TYPE "UDT_Actions"
VERSION : 0.1
   STRUCT
      MCMovement01WP : Bool;   // 1: Fapo in Vorpos AS
      MCMovement02WP : Bool;   // 2: Fapo in AS
      MCMovement03WP : Bool;   // 3: Fapu in Vorpos AS
      MCMovement04WP : Bool;   // 4: Fapu in AS
      MCMovement05WP : Bool;   // 5: Gestell in Vorpos AS
      MCMovement06WP : Bool;   // 6: Gestell in AS
      MCMovement07WP : Bool;   // 7: Parallelhub in Vorpos AS
      MCMovement08WP : Bool;   // 8: Parallelhub in AS
      MCMovement09WP : Bool;   // 9: Parallelhub unten (Fapu mit Fapo) verriegeln
      MCMovement10WP : Bool;   // 10: Sicherheitsriegel Parallelhub entriegeln
      MCMovement11WP : Bool;   // 11: Luftkissen aufblasen
      MCMovement12WP : Bool;   // 12: Form erkannt
      MCMovement13WP : Bool;   // 13: Sicherheitsriegel Fapo entriegeln
      MCMovement14WP : Bool;   // 14: Fapo referenzieren
      MCMovement15WP : Bool;   // 15: Fapu referenzieren
      MCMovement16WP : Bool;   // 16: Gestell referenzieren
      MCMovement17WP : Bool;   // 17: Rolltor zu
      MCMovement18WP : Bool;   // 18: Anschlag Fapo verriegeln
      MCMovement19WP : Bool;   // 19: Sicherheitsriegel Gestell entriegeln
      MCMovement20WP : Bool;   // 20:
      MCMovement21WP : Bool;   // 21:
      MCMovement22WP : Bool;   // 22:
      MCMovement23WP : Bool;   // 23:
      MCMovement24WP : Bool;   // 24:
      MCMovement25WP : Bool;   // 25: Werkzeugriegel Fapo verriegeln
      MCMovement26WP : Bool;   // 26: Werkzeugriegel Fapu verriegeln
      MCMovement27WP : Bool;   // 27: Hubleiste Fapu absenken
      MCMovement28WP : Bool;   // 28: Luftkissen aufblasen (kleiner Druck für Magnet)
      MCMovement29WP : Bool;   // 29: Magnetplatte Fapo einschalten
      MCMovement30WP : Bool;   // 30: Magnetplatte Fapu einschalten
      MCMovement31WP : Bool;   // 31: Fallsicherung Fapo verriegeln
      MCMovement32WP : Bool;   // 32: Fallsicherung Fapu verriegeln
      MCMovement01BP : Bool;   // 33: Fapo in Vorpos GS
      MCMovement02BP : Bool;   // 34: Fapo in GS
      MCMovement03BP : Bool;   // 35: Fapu in Vorpos GS
      MCMovement04BP : Bool;   // 36: Fapu in GS
      MCMovement05BP : Bool;   // 37: Gestell in Vorpos GS
      MCMovement06BP : Bool;   // 38: Gestell in GS
      MCMovement07BP : Bool;   // 39: Parallelhub in Vorpos GS
      MCMovement08BP : Bool;   // 40: Parallelhub in GS
      MCMovement09BP : Bool;   // 41: Parallelhub unten (Fapu mit Fapo) entriegeln
      MCMovement10BP : Bool;   // 42: Sicherheitsriegel Parallelhub verriegeln
      MCMovement11BP : Bool;   // 43: Luftkissen ablassen
      MCMovement12BP : Bool;   // 44:
      MCMovement13BP : Bool;   // 45: Sicherheitsriegel Fapo verriegeln
      MCMovement14BP : Bool;   // 46: Parallelhub in GS od. in Vorpos GS
      MCMovement15BP : Bool;   // 47:
      MCMovement16BP : Bool;   // 48: Parallelhub referenzieren
      MCMovement17BP : Bool;   // 49: Rolltor auf
      MCMovement18BP : Bool;   // 50: Anschlag Fapo entriegeln
      MCMovement19BP : Bool;   // 51: Sicherheitsriegel Gestell verriegeln
      MCMovement20BP : Bool;   // 52:
      MCMovement21BP : Bool;   // 53:
      MCMovement22BP : Bool;   // 54:
      MCMovement23BP : Bool;   // 55:
      MCMovement24BP : Bool;   // 56:
      MCMovement25BP : Bool;   // 57: Werkzeugriegel Fapo entriegeln
      MCMovement26BP : Bool;   // 58: Werkzeugriegel Fapu entriegeln
      MCMovement27BP : Bool;   // 59: Hubleiste Fapu anheben
      MCMovement28BP : Bool;   // 60:
      MCMovement29BP : Bool;   // 61: Magnetplatte Fapo ausschalten
      MCMovement30BP : Bool;   // 62: Magnetplatte Fapu ausschalten
      MCMovement31BP : Bool;   // 63: Fallsicherung Fapo entriegeln
      MCMovement32BP : Bool;   // 64: Fallsicherung Fapu entriegeln
      MouldMovement01WP : Bool;   // 65: Pneumatischer Kernzug DLV-1 ausfahren UT / Hydraulischer Kernzug HV-1
      MouldMovement02WP : Bool;   // 66: Pneumatischer Kernzug DLV-2 ausfahren UT / Hydraulischer Kernzug HV-2
      MouldMovement03WP : Bool;   // 67: Pneumatischer Kernzug DLV-3 ausfahren UT / Hydraulischer Kernzug HV-3
      MouldMovement04WP : Bool;   // 68: Pneumatischer Kernzug DLV-4 ausfahren UT / Hydraulischer Kernzug HV-4
      MouldMovement05WP : Bool;   // 69: Pneumatischer Kernzug DLV-5 ausfahren UT / Hydraulischer Kernzug HV-5
      MouldMovement06WP : Bool;   // 70: Pneumatischer Kernzug DLV-6 ausfahren UT / Hydraulischer Kernzug HV-6
      MouldMovement07WP : Bool;   // 71: Pneumatischer Kernzug DLV-7 ausfahren UT / Pneumatischer Kernzug DLV-1
      MouldMovement08WP : Bool;   // 72: Pneumatischer Kernzug DLV-8 ausfahren UT / Pneumatischer Kernzug DLV-2
      MouldMovement09WP : Bool;   // 73: Pneumatischer Kernzug DLV-1 ausfahren OT / Pneumatischer Kernzug DLV-3
      MouldMovement10WP : Bool;   // 74: Pneumatischer Kernzug DLV-2 ausfahren OT / Pneumatischer Kernzug DLV-4
      MouldMovement11WP : Bool;   // 75: Pneumatischer Kernzug DLV-3 ausfahren OT / Pneumatischer Kernzug DLV-5
      MouldMovement12WP : Bool;   // 76: Pneumatischer Kernzug DLV-4 ausfahren OT / Pneumatischer Kernzug DLV-6
      MouldMovement13WP : Bool;   // 77: Pneumatischer Kernzug DLV-5 ausfahren OT / Pneumatischer Kernzug DLV-7
      MouldMovement14WP : Bool;   // 78: Pneumatischer Kernzug DLV-6 ausfahren OT / Pneumatischer Kernzug DLV-8
      MouldMovement15WP : Bool;   // 79: Pneumatischer Kernzug DLV-7 ausfahren OT
      MouldMovement16WP : Bool;   // 80: Pneumatischer Kernzug DLV-8 ausfahren OT
      MouldMovement17WP : Bool;   // 81:
      MouldMovement18WP : Bool;   // 82:
      MouldMovement19WP : Bool;   // 83:
      MouldMovement20WP : Bool;   // 84:
      MouldMovement21WP : Bool;   // 85:
      MouldMovement22WP : Bool;   // 86:
      MouldMovement23WP : Bool;   // 87:
      MouldMovement24WP : Bool;   // 88: Vakuumventil VV-1 Fapu ansteuern
      MouldMovement25WP : Bool;   // 89: Vakuumventil VV-2 Fapu ansteuern
      MouldMovement26WP : Bool;   // 90: Vakuumventil VV-3 Fapu ansteuern
      MouldMovement27WP : Bool;   // 91: Vakuumventil VV-1 Fapo ansteuern
      MouldMovement28WP : Bool;   // 92: Vakuumventil VV-2 Fapo ansteuern
      MouldMovement29WP : Bool;   // 93: Vakuumventil VV-3 Fapo ansteuern
      MouldMovement30WP : Bool;   // 94: Vakuumtest VV-1 Fapu
      MouldMovement31WP : Bool;   // 95: Vakuumtest VV-2 Fapu
      MouldMovement32WP : Bool;   // 96: Vakuumtest VV-3 Fapu
      MouldMovement01BP : Bool;   // 97: Pneumatischer Kernzug DLV-1 einfahren UT / Hydraulischer Kernzug HV-1
      MouldMovement02BP : Bool;   // 98: Pneumatischer Kernzug DLV-2 einfahren UT / Hydraulischer Kernzug HV-2
      MouldMovement03BP : Bool;   // 99: Pneumatischer Kernzug DLV-3 einfahren UT / Hydraulischer Kernzug HV-3
      MouldMovement04BP : Bool;   // 100: Pneumatischer Kernzug DLV-4 einfahren UT / Hydraulischer Kernzug HV-4
      MouldMovement05BP : Bool;   // 101: Pneumatischer Kernzug DLV-5 einfahren UT / Hydraulischer Kernzug HV-5
      MouldMovement06BP : Bool;   // 102: Pneumatischer Kernzug DLV-6 einfahren UT / Hydraulischer Kernzug HV-6
      MouldMovement07BP : Bool;   // 103: Pneumatischer Kernzug DLV-7 einfahren UT / Pneumatischer Kernzug DLV-1
      MouldMovement08BP : Bool;   // 104: Pneumatischer Kernzug DLV-8 einfahren UT / Pneumatischer Kernzug DLV-2
      MouldMovement09BP : Bool;   // 105: Pneumatischer Kernzug DLV-1 einfahren OT / Pneumatischer Kernzug DLV-3
      MouldMovement10BP : Bool;   // 106: Pneumatischer Kernzug DLV-2 einfahren OT / Pneumatischer Kernzug DLV-4
      MouldMovement11BP : Bool;   // 107: Pneumatischer Kernzug DLV-3 einfahren OT / Pneumatischer Kernzug DLV-5
      MouldMovement12BP : Bool;   // 108: Pneumatischer Kernzug DLV-4 einfahren OT / Pneumatischer Kernzug DLV-6
      MouldMovement13BP : Bool;   // 109: Pneumatischer Kernzug DLV-5 einfahren OT / Pneumatischer Kernzug DLV-7
      MouldMovement14BP : Bool;   // 110: Pneumatischer Kernzug DLV-6 einfahren OT / Pneumatischer Kernzug DLV-8
      MouldMovement15BP : Bool;   // 111: Pneumatischer Kernzug DLV-7 einfahren OT
      MouldMovement16BP : Bool;   // 112: Pneumatischer Kernzug DLV-8 einfahren OT
      MouldMovement17BP : Bool;   // 113:
      MouldMovement18BP : Bool;   // 114:
      MouldMovement19BP : Bool;   // 115:
      MouldMovement20BP : Bool;   // 116:
      MouldMovement21BP : Bool;   // 117:
      MouldMovement22BP : Bool;   // 118:
      MouldMovement23BP : Bool;   // 119:
      MouldMovement24BP : Bool;   // 120: Vakuumventil VV-1 Fapu absteuern
      MouldMovement25BP : Bool;   // 121: Vakuumventil VV-2 Fapu absteuern
      MouldMovement26BP : Bool;   // 122: Vakuumventil VV-3 Fapu absteuern
      MouldMovement27BP : Bool;   // 123: Vakuumventil VV-1 Fapo absteuern
      MouldMovement28BP : Bool;   // 124: Vakuumventil VV-2 Fapo absteuern
      MouldMovement29BP : Bool;   // 125: Vakuumventil VV-3 Fapo absteuern
      MouldMovement30BP : Bool;   // 126: Vakuumtest VV-1 Fapo
      MouldMovement31BP : Bool;   // 127: Vakuumtest VV-2 Fapo
      MouldMovement32BP : Bool;   // 128: Vakuumtest VV-3 Fapo
      ShotPreparation : Bool;   // 129: Schussvorbereitung ausgeben
      ShotEnable : Bool;   // 130: Schussfreigabe ausgeben
      ShotEnd : Bool;   // 131: Schussende abwarten
      StartReactionTime : Bool;   // 132: Reaktionszeit starten
      WaitReactionTime : Bool;   // 133: Reaktionszeit abwarten
      Spare134 : Bool;   // 134:
      Spare135 : Bool;   // 135:
      Spare136 : Bool;   // 136:
      Spare137 : Bool;   // 137:
      Spare138 : Bool;   // 138:
      WaitTime1 : Bool;   // 139: Ablauf der Wartezeit 1
      WaitTime2 : Bool;   // 140: Ablauf der Wartezeit 2
      WaitTime3 : Bool;   // 141: Ablauf der Wartezeit 3
      WaitTime4 : Bool;   // 142: Ablauf der Wartezeit 4
      WaitTime5 : Bool;   // 143: Ablauf der Wartezeit 5
      WaitTime6 : Bool;   // 144: Ablauf der Wartezeit 6
      StopCycle : Bool;   // 145: Zyklus unterbrechen
      Spare146 : Bool;   // 146:
      NoFaultGroup1 : Bool;   // 147: Keine Sörgruppe 1
      SafetyOk : Bool;   // 148: Sicherheit ok
      StartWatch : Bool;   // 149: Start Stoppuhr
      StopWatch : Bool;   // 150: Stop Stoppuhr
      Spare151 : Bool;   // 151:
      Spare152 : Bool;   // 152:
      Spare153 : Bool;   // 153:
      Spare154 : Bool;   // 154:
      Spare155 : Bool;   // 155:
      Spare156 : Bool;   // 156:
      Set_access_release : Bool;   // 157: Zutrittsfreigabe setzen
      Reset_access_release : Bool;   // 158: Zutrittsfreigabe zurücksetzen
      RobotOutOfMC : Bool;   // 159: Roboter nicht im Bereich des Formträgers
      EndOfProgram : Bool;   // 160: Programm Ende
   END_STRUCT;
END_TYPE

TYPE "UDT_CoreSettings"
VERSION : 0.1
   STRUCT
      Bit_Inverted_WP_01 : Bool;
      Bit_inverted_WP_02 : Bool;
      Bit_inverted_WP_03 : Bool;
      Bit_inverted_WP_04 : Bool;
      Bit_inverted_WP_05 : Bool;
      Bit_inverted_WP_06 : Bool;
      Signal_from_upper_tool_WP : Bool;
      Always_ON_WP : Bool;
      Bit_inverted_BP_01 : Bool;
      Bit_inverted_BP_02 : Bool;
      Bit_inverted_BP_03 : Bool;
      Bit_inverted_BP_04 : Bool;
      Bit_inverted_BP_05 : Bool;
      Bit_inverted_BP_06 : Bool;
      Signal_from_upper_tool_BP : Bool;
      Always_ON_BP : Bool;
      Pin_No_WP_01 : Int;
      Pin_No_WP_02 : Int;
      Pin_No_WP_03 : Int;
      Pin_No_WP_04 : Int;
      Pin_No_WP_05 : Int;
      Pin_No_WP_06 : Int;
      Spare_14 : Int;
      Pin_No_BP_01 : Int;
      Pin_No_BP_02 : Int;
      Pin_No_BP_03 : Int;
      Pin_No_BP_04 : Int;
      Pin_No_BP_05 : Int;
      Pin_No_BP_06 : Int;
      Spare_28 : Int;
   END_STRUCT;
END_TYPE

TYPE "UDT_CoreSettingsSpecial"
VERSION : 0.1
   STRUCT
      EndPos_Byte_WP_1 : Byte;   // Eingangsbyte für die Endposition
      EndPos_Byte_WP_2 : Byte;   // Eingangsbyte für die Endposition
      EndPos_Byte_WP_3 : Byte;   // Eingangsbyte für die Endposition
      EndPos_Byte_WP_4 : Byte;   // Eingangsbyte für die Endposition
      EndPos_Byte_WP_5 : Byte;   // Eingangsbyte für die Endposition
      EndPos_Byte_WP_6 : Byte;   // Eingangsbyte für die Endposition
      EndPos_Bit_WP_1 : Byte;   // Eingangsbyte für die Endposition
      EndPos_Bit_WP_2 : Byte;   // Eingangsbyte für die Endposition
      EndPos_Bit_WP_3 : Byte;   // Eingangsbyte für die Endposition
      EndPos_Bit_WP_4 : Byte;   // Eingangsbyte für die Endposition
      EndPos_Bit_WP_5 : Byte;   // Eingangsbyte für die Endposition
      EndPos_Bit_WP_6 : Byte;   // Eingangsbyte für die Endposition
      EndPos_Byte_BP_1 : Byte;   // Eingangsbyte für die Endposition
      EndPos_Byte_BP_2 : Byte;   // Eingangsbyte für die Endposition
      EndPos_Byte_BP_3 : Byte;   // Eingangsbyte für die Endposition
      EndPos_Byte_BP_4 : Byte;   // Eingangsbyte für die Endposition
      EndPos_Byte_BP_5 : Byte;   // Eingangsbyte für die Endposition
      EndPos_Byte_BP_6 : Byte;   // Eingangsbyte für die Endposition
      EndPos_Bit_BP_1 : Byte;   // Eingangsbyte für die Endposition
      EndPos_Bit_BP_2 : Byte;   // Eingangsbyte für die Endposition
      EndPos_Bit_BP_3 : Byte;   // Eingangsbyte für die Endposition
      EndPos_Bit_BP_4 : Byte;   // Eingangsbyte für die Endposition
      EndPos_Bit_BP_5 : Byte;   // Eingangsbyte für die Endposition
      EndPos_Bit_BP_6 : Byte;   // Eingangsbyte für die Endposition
   END_STRUCT;
END_TYPE

TYPE "UDT_Limit_axis"
VERSION : 0.1
   STRUCT
      Speed_manual : Struct
         VPosWP : Int;
         VPrePosWP : Int;
         VPrePosBP : Int;
         VPosBP : Int;
      END_STRUCT;
      Speed_auto : Struct
         VPosWP : Int;
         VPrePosWP : Int;
         VPrePosBP : Int;
         VPosBP : Int;
      END_STRUCT;
      Acceleration : Struct
         Min_value : Struct
            PosWP : Int;
            PrePosWP : Int;
            PrePosBP : Int;
            PosBP : Int;
         END_STRUCT;
         Max_value : Struct
            PosWP : Int;
            PrePosWP : Int;
            PrePosBP : Int;
            PosBP : Int;
         END_STRUCT;
      END_STRUCT;
      Deceleration : Struct
         Min_value : Struct
            PosWP : Int;
            PrePosWP : Int;
            PrePosBP : Int;
            PosBP : Int;
         END_STRUCT;
         Max_value : Struct
            PosWP : Int;
            PrePosWP : Int;
            PrePosBP : Int;
            PosBP : Int;
         END_STRUCT;
      END_STRUCT;
      Movement : Struct
         Min_value : Struct
            PosWP : Real;
            PrePosWP : Real;
            PrePosBP : Real;
            PosBP : Real;
         END_STRUCT;
         Max_value : Struct
            PosWP : Real;
            PrePosWP : Real;
            PrePosBP : Real;
            PosBP : Real;
         END_STRUCT;
      END_STRUCT;
      Switch_over_pos : Struct
         Start : Struct
            PosWP : Real;
            PrePosWP : Real;
            PrePosBP : Real;
            PosBP : Real;
         END_STRUCT;
         End : Struct
            PosWP : Real;
            PrePosWP : Real;
            PrePosBP : Real;
            PosBP : Real;
         END_STRUCT;
      END_STRUCT;
   END_STRUCT;
END_TYPE

TYPE "UDT_TempPulse"
VERSION : 0.1
   STRUCT
      Wichtung : Int := 0;
      MaxDelta_K : Int := 0;
      MaxDelta_H : Int := 0;
      Min_Time : Int := 0;
      Regelstrecke : Int := 0;
      Bits : Struct
         Start_TON : Bool;
         Status_TON : Bool;
      END_STRUCT;
      Heizen : Bool := FALSE;
      Kuehlen : Bool := FALSE;
      Reserve : Bool := FALSE;
      Reserve1 : Bool := FALSE;
      Reserve3 : Bool := FALSE;
      Reserve4 : Bool := FALSE;
      Reserve5 : Bool := FALSE;
      Reserve6 : Bool := FALSE;
   END_STRUCT;
END_TYPE

TYPE "UDT071_CPiston_State"
TITLE = State of cleaning piston at mixing head
VERSION : 0.0
   STRUCT
      FaultLevel_1 : Bool;
      FaultLevel_2 : Bool;
      FaultLevel_3 : Bool;
      FaultExists : Bool;
      Edge_MH_was_open : Bool;   // Edge flag to detect mixinghead was open
      PS_not_released : Bool;   // Partshot is blocked (like service shot)
      Edge_CP_nOK : Bool;   // Edge flag to delete signal "IO_CP_is_ok" of foaming release
      CP_is_OK : Bool;   // Activation of cleaning piston is ok (like signal "IO_RK_is_ok")
      MH_was_open : Bool;   // Information cleanig necessary, because mixing head was open
      Switch_CP_Forward : Bool;   // Cleaning stroke forward
      CleanAfterShotSelected : Bool;   // Cleaning of mixinghead is requested after part shot
      CleaningFromEPrunning : Bool;   // Cleaning stroke request from external plant is running
      Cleaning_runs : Bool;   // General information cleaning stroke active
      Spare_1_5 : Bool;
      CP_Moved_Manual : Bool;   // The cleaning CP was moved manual
      CP_valve_selected : Bool;   // Activation of valve cleaning from cleaning piston is selected
      Stop_Cleaning : Bool;   // Information cleanig stroke cleanig piston finished
      Stepnumber : Byte;   // Stepnumber of steps sequence control cleaning piston
      State_CP : Byte;   // 1->CP Forward; 2->Fault CP; 3->CP requested but not on
   END_STRUCT;
END_TYPE

TYPE "UDT_CorePosition_Special"
VERSION : 0.1
   STRUCT
      EndPos_WP_1 : Bool;   // Endlage erreicht
      EndPos_WP_2 : Bool;   // Endlage erreicht
      EndPos_WP_3 : Bool;   // Endlage erreicht
      EndPos_WP_4 : Bool;   // Endlage erreicht
      EndPos_WP_5 : Bool;   // Endlage erreicht
      EndPos_WP_6 : Bool;   // Endlage erreicht
      Spare_0_6 : Bool;
      Spare_0_7 : Bool;
      EndPos_BP_1 : Bool;   // Endlage erreicht
      EndPos_BP_2 : Bool;   // Endlage erreicht
      EndPos_BP_3 : Bool;   // Endlage erreicht
      EndPos_BP_4 : Bool;   // Endlage erreicht
      EndPos_BP_5 : Bool;   // Endlage erreicht
      EndPos_BP_6 : Bool;   // Endlage erreicht
      Spare_1_6 : Bool;
      Spare_1_7 : Bool;
   END_STRUCT;
END_TYPE

TYPE "UDT073_CP_StateMQMX"
VERSION : 0.0
   STRUCT
      Stoer_LFZRKVor_MQ : Bool;
      Stoer_LFZRKZurueck_MQ : Bool;
      Stoer_LFZDrosselVor_MQ : Bool;
      Stoer_LFZDrossZurueck_MQ : Bool;
      Stoer_Dosierstellung_MQ : Bool;
      Stoer_Grundstellung_MQ : Bool;
      Stoer_Initiatoren_MQ : Bool;
      Stoer_LFZRK_MX : Bool;
      Stoer_LFZDrossel_MX : Bool;
      Stoer_LFZDosierkolben_MX : Bool;
      Stoer_Dosierstellung_MX : Bool;
      Res_STG1 : Bool;
      Res_STG2 : Bool;
      Res_STG3 : Bool;
      Res_STG4 : Bool;
      Reinigungskolben_Ok : Bool;
      Anforderung_von_RK : Bool;
      WartezReinigenLaeuft : Bool;
      ReinigenLaeuft : Bool;
      WartezTaktLaeuft : Bool;
      TaktreinigenLAeuft : Bool;
      Handreinigen : Bool;
      ReinigenNachDosieren : Bool;
      ReinigungstaktLaeuft : Bool;
      WartenAufRK : Bool;
      ReinigenEIN : Bool;
      Reserve2 : Bool;
      Reserve3 : Bool;
      VW_Einzelbewegung_RK : Bool;
      VW_Einzelbewegung_Dross : Bool;
      VW_Intervallreinigung : Bool;
      VW_Ini_Dosierkolben_Brue : Bool;
      VFZ_Drosselschieber : S5Time := S5T#800MS;
      VFZ_Reinigungskolben : S5Time := S5T#2S;
      VFZ_DrosselvorKolben : S5Time := S5T#1S;
      WartezeitReinigen : S5Time := S5T#500MS;
      Reinigungszeit : S5Time := S5T#20S;
      WartezeitIntervallrein : S5Time := S5T#10S;
      ReinigungszeitIntervall : S5Time := S5T#50S;
      ReinigenIntervallfolgez : S5Time := S5T#8S;
      Reserve_T1 : S5Time;
      Reserve_T2 : S5Time;
      Reserve_T3 : S5Time;
      Reserve_T4 : S5Time;
      Reserve_T5 : S5Time;
   END_STRUCT;
END_TYPE

TYPE "UDT_ET200SP_config"
VERSION : 0.1
   STRUCT
      Block_length : Byte := 20;   // 4+(2*number of slots)
      Block_ID : Byte := 196;   // Data record number
      "Version" : Byte := 2;
      Subversion : Byte := 0;
      Card : Array[1..8] of Struct
         slot : Byte;   // configured slot 1 < real slot
         add : Byte;   // additional function slot
      END_STRUCT;
   END_STRUCT;
   // Card[1].slot := 16#1;
   // Card[1].add := 0;
   // Card[2].slot := 16#2;
   // Card[3].slot := 16#3;
   // Card[4].slot := 16#4;
   // Card[5].slot := 16#5;
   // Card[6].slot := 16#6;
   // Card[7].slot := 16#7;
   // Card[7].add := 0;
   // Card[6].add := 0;
   // Card[5].add := 0;
   // Card[4].add := 0;
   // Card[3].add := 0;
   // Card[2].add := 0;
END_TYPE

TYPE "UDT_Tool_Outputs_type_1"
VERSION : 0.1
   STRUCT
      "Lower Mould" : Struct
         "2A4" : Struct
            O_Vacuum_WS : Bool := FALSE;   // 0.0
            O_Vacuum_Cavity : Bool := FALSE;   // 0.1
            O_Vacuum_Run_OFF : Bool := FALSE;   // 0.2
            Element_1 : Bool := FALSE;   // 0.3
            Element_2 : Bool := FALSE;   // 0.4
            O_Vacuum_ventilate : Bool := FALSE;   // 0.5
            Element_3 : Bool := FALSE;   // 0.6
            Element_4 : Bool := FALSE;   // 0.7
            Element_5 : Bool := FALSE;   // 1.0
            Element_6 : Bool := FALSE;   // 1.1
            O_Seal_01 : Bool := FALSE;   // 1.2
            O_Seal_02 : Bool := FALSE;   // 1.3
            O_Seal_03 : Bool := FALSE;   // 1.4
            O_Seal_04 : Bool := FALSE;   // 1.5
            O_Seal_05 : Bool := FALSE;   // 1.6
            O_Seal_06 : Bool := FALSE;   // 1.7
         END_STRUCT;
         "2A5" : Struct
            O_Seal_07 : Bool := FALSE;   // 0.0
            O_Seal_08 : Bool := FALSE;   // 0.1
            O_Seal_09 : Bool := FALSE;   // 0.2
            O_Seal_10 : Bool := FALSE;   // 0.3
            O_Seal_11 : Bool := FALSE;   // 0.4
            O_Seal_12 : Bool := FALSE;   // 0.5
            O_Seal_13 : Bool := FALSE;   // 0.6
            O_Seal_14 : Bool := FALSE;   // 0.7
            Element_1 : Bool := FALSE;   // 1.0
            O_LED_Vacuum_WS : Bool := FALSE;   // 1.1
            O_LED_Vacuum_Cavity : Bool := FALSE;   // 1.2
            O_LED_Vacuum_Run_off : Bool := FALSE;   // 1.3
            Element_4 : Bool := FALSE;   // 1.4
            Element_6 : Bool := FALSE;   // 1.5
            Element_7 : Bool := FALSE;   // 1.6
            O_Valve_Seal_on_6Bar : Bool := FALSE;   // 1.7
         END_STRUCT;
         "2A6" : Struct
            O_LED_Sensor_upper_part_substrate_detect : Bool := FALSE;   // 0.0
            O_LED_Sensor_upper_part_substrate_flamed : Bool := FALSE;   // 0.1
            O_LED_Sensor_upper_part_substrate_additionalpart : Bool := FALSE;   // 0.2
            O_LED_Sensor_upper_part_Airbag_WP : Bool := FALSE;   // 0.3
            O_LED_Sensor_lower_part_vacuum_WP : Bool := FALSE;   // 0.4
            O_Pusher_Sealing_WP : Bool := FALSE;   // 0.5
            O_Pusher_Sealing_BP : Bool := FALSE;   // 0.6
            O_Ejector_BP : Bool := FALSE;   // 0.7
            Element_2 : Bool := FALSE;   // 1.0
            Element_3 : Bool := FALSE;   // 1.1
            Element_4 : Bool := FALSE;   // 1.2
            Element_5 : Bool := FALSE;   // 1.3
            Element_6 : Bool := FALSE;   // 1.4
            Element_7 : Bool := FALSE;   // 1.5
            Element_8 : Bool := FALSE;   // 1.6
            Element_9 : Bool := FALSE;   // 1.7
         END_STRUCT;
         "2A8" : Struct
            O_Pusher_Windshield_WP : Bool := FALSE;   // 0.0
            O_Pusher_Windshield_BP : Bool := FALSE;   // 0.1
            O_Pusher_Knee_Border_WP : Bool := FALSE;   // 0.2
            O_Pusher_Knee_Border_BP : Bool := FALSE;   // 0.3
            O_Pusher_Frontal_Area_WP : Bool := FALSE;   // 0.4
            O_Pusher_Frontal_Area_BP : Bool := FALSE;   // 0.5
            O_Ejector_WP : Bool := FALSE;   // 0.6
            Element_1 : Bool := FALSE;   // 0.7
            O_Pusher_Stössel_WP : Bool := FALSE;   // 1.0
            O_Pusher_Stössel_BP : Bool := FALSE;   // 1.1
            O_Flip_Flap_Knee_WP : Bool := FALSE;   // 1.2
            O_Flip_Flap_Knee_BP : Bool := FALSE;   // 1.3
            O_Pusher_Savtey_locking_Knee_WP : Bool := FALSE;   // 1.4
            O_Pusher_Savtey_locking_Knee_BP : Bool := FALSE;   // 1.5
            O_Pusher_Savtey_locking_WS_WP : Bool := FALSE;   // 1.6
            O_Pusher_Savtey_locking_WS_BP : Bool := FALSE;   // 1.7
         END_STRUCT;
         "2A9" : Struct
            O_Pusher_circuit_breakers_WP_SET : Bool := FALSE;   // 0.0
            O_Pusher_circuit_breakers_WP_CLR : Bool := FALSE;   // 0.1
            O_Pusher_circuit_breakers_BP_SET : Bool := FALSE;   // 0.2
            O_Pusher_circuit_breakers_BP_CLR : Bool := FALSE;   // 0.3
            Element_5 : Bool := FALSE;   // 0.4
            Element_6 : Bool := FALSE;   // 0.5
            Element_7 : Bool := FALSE;   // 0.6
            Element_8 : Bool := FALSE;   // 0.7
            Element_1 : Bool := FALSE;   // 1.0
            Element_2 : Bool := FALSE;   // 1.1
            Element_9 : Bool := FALSE;   // 1.2
            Element_10 : Bool := FALSE;   // 1.3
            Element_11 : Bool := FALSE;   // 1.4
            Element_12 : Bool := FALSE;   // 1.5
            Element_13 : Bool := FALSE;   // 1.6
            Element_14 : Bool := FALSE;   // 1.7
         END_STRUCT;
      END_STRUCT;
      "Upper Mould" : Struct
         "46A2" : Struct
            Element_1 : Bool := FALSE;   // 0.0
            O_Pusher_Airbag_BP : Bool := FALSE;   // 0.1
            O_Vacuum_Cups_on : Bool := FALSE;   // 0.2
            O_Vacuum_cavity_on : Bool := FALSE;   // 0.3
            O_Vacuum_ventilate : Bool := FALSE;   // 0.4
            Reserve_5 : Bool := FALSE;   // 0.5
            Reserve_6 : Bool := FALSE;   // 0.6
            O_Indicator_Lamp_Vacuum_on : Bool := FALSE;   // 0.7
            Reserve_13 : Bool := FALSE;   // 1.0
            Reserve_12 : Bool := FALSE;   // 1.1
            Reserve_11 : Bool := FALSE;   // 1.2
            Reserve_10 : Bool := FALSE;   // 1.3
            Reserve_9 : Bool := FALSE;   // 1.4
            Reserve_8 : Bool := FALSE;   // 1.5
            Reserve_7 : Bool := FALSE;   // 1.6
            Reserve_14 : Bool := FALSE;   // 1.7
         END_STRUCT;
         "46A4" : Struct
            O_Pusher_Airbag_WP : Bool := FALSE;   // 0.0
            Element_1 : Bool := FALSE;   // 0.1
            O_Pusher_WP : Bool := FALSE;   // 0.2
            O_Pusher_BP : Bool := FALSE;   // 0.3
            Reserve_12 : Bool := FALSE;   // 0.4
            Reserve_13 : Bool := FALSE;   // 0.5
            Reserve_14 : Bool := FALSE;   // 0.6
            Reserve_15 : Bool := FALSE;   // 0.7
            Reserve_16 : Bool := FALSE;   // 1.0
            Reserve_17 : Bool := FALSE;   // 1.1
            Reserve_11 : Bool := FALSE;   // 1.2
            Reserve_10 : Bool := FALSE;   // 1.3
            Reserve_9 : Bool := FALSE;   // 1.4
            Reserve_8 : Bool := FALSE;   // 1.5
            Reserve_7 : Bool := FALSE;   // 1.6
            Reserve_18 : Bool := FALSE;   // 1.7
         END_STRUCT;
      END_STRUCT;
   END_STRUCT;
END_TYPE

TYPE "UDT_Word_1-16"
VERSION : 0.1
   STRUCT
      "01" : Bool;
      "02" : Bool;
      "03" : Bool;
      "04" : Bool;
      "05" : Bool;
      "06" : Bool;
      "07" : Bool;
      "08" : Bool;
      "09" : Bool;
      "10" : Bool;
      "11" : Bool;
      "12" : Bool;
      "13" : Bool;
      "14" : Bool;
      "15" : Bool;
      "16" : Bool;
      "17" : Bool;
      "18" : Bool;
      "19" : Bool;
      "20" : Bool;
      "21" : Bool;
      "22" : Bool;
      "23" : Bool;
      "24" : Bool;
      "25" : Bool;
      "26" : Bool;
      "27" : Bool;
      "28" : Bool;
      "29" : Bool;
      "30" : Bool;
      "31" : Bool;
      "32" : Bool;
   END_STRUCT;
END_TYPE

TYPE "UDT_Siemens_FC"
VERSION : 0.1
   STRUCT
      HW_ID : Hw_Any;
      Input : Struct
         Schleppabstand_in_Toleranz : Bool;
         Führung_gefordert : Bool;
         Zielposition_erreicht : Bool;
         Referenzpunkt_gesetzt : Bool;
         Quittierung_Verfahrsatz_aktiviert : Bool;
         Drehzahlschwellwert : Bool;
         Achse_beschleunigt : Bool;
         Achse_verzögert : Bool;
         Einschaltbereit : Bool;
         Betriebsbereit : Bool;
         Ready_to_run : Bool;
         Störung_wirksam : Bool;
         Kein_Austrudeln_aktiv : Bool;
         Kein_Schnellhalt_aktiv : Bool;
         Einschaltsperre_aktiv : Bool;
         Warnung_wirksam : Bool;
         "15" : Bool;
         "16" : Bool;
         "17" : Bool;
         "18" : Bool;
         "19" : Bool;
         Profil_aktiv : Bool;
         "21" : Bool;
         MDI_aktiv : Bool;
      END_STRUCT;
   END_STRUCT;
END_TYPE

TYPE "UDT_OperatingMode"
VERSION : 0.1
   STRUCT
      valid : Bool;
      manual : Bool;
      semi_automatic : Bool;
      automatic : Bool;
      control_voltage : Bool;
      HF_manual : Bool;
      Pulse_manual : Bool;
      HF_semi_automatic : Bool;
      Pulse_semi_automatic : Bool;
      FH_automatic : Bool;
      Pulse_automatic : Bool;
      HF_request_start : Bool;
      Request_start : Bool;
      HF_OM_0 : Bool;
      Pulse_OM_0 : Bool;
      Automatic_stop_okay : Bool;
      Lamp_test : Bool;
      Start_production : Bool;
      Production : Bool;
      Stop_production : Bool;
      Button_semic_automatic : Bool;
      Semi_automatic_active : Bool;
      Alarm_active : Bool;   // Alarm aktiv an OP
      Reference : Bool;
      Operating_mode_to_TP : Byte;   // 1: Control voltage; 2: manual; 3: automatik; 4: Cycle running
   END_STRUCT;
END_TYPE

TYPE "UDT_Mould_status"
VERSION : 0.1
   STRUCT
      HM_OT_1 : Bool;
      HM_OT_2 : Bool;
      HM_OT_3 : Bool;
      HM_OT_4 : Bool;
      HM_OT_5 : Bool;
      HM_OT_6 : Bool;
      HM_OT_7 : Bool;
      HM_OT_8 : Bool;
      HM_UT_1 : Bool;
      HM_UT_2 : Bool;
      HM_UT_3 : Bool;
      HM_UT_4 : Bool;
      HM_UT_5 : Bool;
      HM_UT_6 : Bool;
      HM_UT_7 : Bool;
      HM_UT_8 : Bool;
      M_UT_auf : Bool;
      FHM_2Hand : Bool;
      HM_SchieberSichern_1 : Bool;
      HM_SchieberSichern_2 : Bool;
      HM_SchieberSichern_3 : Bool;
      HM_SchieberSichern_4 : Bool;
      HM_SchieberSichern_5 : Bool;
      HM_SchieberSichern_6 : Bool;
      Free_Bit_01 : Bool;
      Free_Bit_02 : Bool;
      Free_Bit_03 : Bool;
      Free_Bit_04 : Bool;
      Free_Bit_05 : Bool;
      Free_Bit_06 : Bool;
      Free_Bit_07 : Bool;
      Free_Bit_08 : Bool;
      Free_Bit_09 : Bool;
      Free_Bit_10 : Bool;
      Free_Bit_11 : Bool;
      Free_Bit_12 : Bool;
      Free_Bit_13 : Bool;
      Free_Bit_14 : Bool;
      Free_Bit_15 : Bool;
      Free_Bit_16 : Bool;
      Free_Byte_01 : Bool;
      Free_Byte_02 : Bool;
      Free_Byte_03 : Bool;
      Free_Byte_04 : Bool;
   END_STRUCT;
END_TYPE

TYPE "UDT_SafetyDevice"
VERSION : 0.1
   STRUCT
      OpeningSelected : Bool;   // Opening of the safety device is selected
      OpeningEnabled : Bool;   // Opening of the safety device is possible
      EdgeButton : Bool;   // Edge of the button to select opening of the safety device
      HFEdgeButton : Bool;   // Help flag for the edge
      EdgeASReset : Bool;   // Edgo of the reset of Auto Stop from this safety device
      HFEdgeASReset : Bool;   // Help flag for the edge
      HFforMESSelected : Bool;   // Help flag for the message opening is selected
      HFforMESAutomaticStop : Bool;   // Help flag for message automatic stop is activ
      Spare_1 : Byte;
      Msg_Selected : Bool;   // Message safety device is selected
      Msg_AS_active : Bool;   // Message autostop from safety device is active
      Spare_2_2 : Bool;
      Spare_2_3 : Bool;
      Spare_2_4 : Bool;
      Spare_2_5 : Bool;
      Spare_2_6 : Bool;
      Spare_2_7 : Bool;
      Spare_3 : Byte;
   END_STRUCT;
END_TYPE

TYPE "UDT_Times_temperatures_tool"
VERSION : 0.1
   STRUCT
      Set_times : Struct   // general use
         Reaction_time_1 : Time := T#1M;
         Reaction_time_2 : Time := T#0MS;
         Reaction_time_3 : Time := T#0MS;
         Reaction_time_4 : Time := T#0MS;
         Reaction_time_5 : Time := T#0MS;
         Reaction_time_6 : Time := T#0MS;
         Time_befor_degasing_tool_1 : Time := T#20S;
         Degasing_time_tool_1 : Time := T#10S;
         Time_befor_degasing_tool_2 : Time := T#0MS;
         Degasing_time_tool_2 : Time := T#0MS;
         Time_befor_degasing_tool_3 : Time := T#0MS;
         Degasing_time_tool_3 : Time := T#0MS;
         Time_befor_degasing_tool_4 : Time := T#0MS;
         Degasing_time_tool_4 : Time := T#0MS;
         Time_befor_degasing_tool_5 : Time := T#0MS;
         Degasing_time_tool_5 : Time := T#0MS;
         Time_befor_degasing_tool_6 : Time := T#0MS;
         Degasing_time_tool_6 : Time := T#0MS;
         Waiting_time_1 : Time := T#10S;
         Waiting_time_2 : Time := T#2S;
         Waiting_time_3 : Time := T#3S;
         Waiting_time_4 : Time := T#4S;
         Waiting_time_5 : Time := T#5S;
         Waiting_time_6 : Time := T#6S;
         Test_vacuum_circit_1 : Time := T#0MS;   // Dauer des Vakuumtestes für den Vakuumkreis 01
         Test_vacuum_circit_2 : Time := T#0MS;   // Dauer des Vakuumtestes für den Vakuumkreis 02
         Test_vacuum_circit_3 : Time := T#0MS;   // Dauer des Vakuumtestes für den Vakuumkreis 03
         Test_vacuum_circit_4 : Time := T#0MS;   // Dauer des Vakuumtestes für den Vakuumkreis 04
         Test_vacuum_circit_5 : Time := T#0MS;   // Dauer des Vakuumtestes für den Vakuumkreis 05
         Test_vacuum_circit_6 : Time := T#0MS;   // Dauer des Vakuumtestes für den Vakuumkreis 06
         Release_vacuum : Time := T#0MS;
         Switch_off_delay_vacuum_pump : Time := T#10S;   // switch off delay for vacuum pump
         Switch_off_delay_exhaust : Time := T#10S;   // Ausschaltverzögerung Klappe Absaugung
         Stopwatch : Time := T#0MS;
         Spare_35 : Time := T#0MS;
         Spare_36 : Time := T#0MS;
         Spare_37 : Time := T#0MS;
         Spare_38 : Time := T#0MS;
         Spare_39 : Time := T#0MS;
         Spare_40 : Time := T#0MS;
         Spare_41 : Time := T#0MS;
         Spare_42 : Time := T#0MS;
         Spare_43 : Time := T#0MS;
      END_STRUCT;
      Set_times_movement : Struct   // running times
         Time_MC_WP : Array[0..32] of Time;
         Time_MC_BP : Array[0..32] of Time;
         Time_MLD_WP : Array[0..32] of Time;
         Time_MLD_BP : Array[0..32] of Time;
      END_STRUCT;
      Set_times_seals : Struct   // seal times
         SOD_seal : Array[0..32] of Time;   // switch on delay seal
         Duration_seal : Array[0..32] of Time;   // duration seal
      END_STRUCT;
      Set_temperature : Struct   // temperature handling
         Setvalue : Array[0..16] of Int;
         Warning_Tolerance : Struct
            Warning_min : Array[0..16] of Int;
            Warning_max : Array[0..16] of Int;
            Tolerance_min : Array[0..16] of Int;
            Tolerance_max : Array[0..16] of Int;
         END_STRUCT;
         Settings_Pulse : Struct
            PulseTemp_K1 : "UDT_TempPulse";
            Pulsezeit_K1 : DInt := 50000;
            PulseTemp_K2 : "UDT_TempPulse";
            Pulsezeit_K2 : DInt := -41943050;
            PulseTemp_K3 : "UDT_TempPulse";
            Pulsezeit_K3 : DInt := 50000;
            PulseTemp_K4 : "UDT_TempPulse";
            Pulsezeit_K4 : DInt := -41943050;
            PulseTemp_K5 : "UDT_TempPulse";
            Pulsezeit_K5 : DInt := -41943050;
            PulseTemp_K6 : "UDT_TempPulse";
            Pulsezeit_K6 : DInt := -41943050;
            PulseTemp_K7 : "UDT_TempPulse";
            Pulsezeit_K7 : DInt := -41943050;
            PulseTemp_K8 : "UDT_TempPulse";
            Pulsezeit_K8 : DInt := -41943050;
            PulseTemp_K9 : "UDT_TempPulse";
            Pulsezeit_K9 : DInt := -41943050;
            PulseTemp_K10 : "UDT_TempPulse";
            Pulsezeit_K10 : DInt := -41943050;
            PulseTemp_K11 : "UDT_TempPulse";
            Pulsezeit_K11 : DInt := -41943050;
            PulseTemp_K12 : "UDT_TempPulse";
            Pulsezeit_K12 : DInt := -41943050;
            PulseTemp_K13 : "UDT_TempPulse";
            Pulsezeit_K13 : DInt := -41943050;
            PulseTemp_K14 : "UDT_TempPulse";
            Pulsezeit_K14 : DInt := -41943050;
            PulseTemp_K15 : "UDT_TempPulse";
            Pulsezeit_K15 : DInt := -41943050;
            PulseTemp_K16 : "UDT_TempPulse";
            Pulsezeit_K16 : DInt := -41943050;
         END_STRUCT;
         Exist : Array[0..16] of Bool;
      END_STRUCT;
      Set_Core_settings : Struct   // core settings WinCap
         Special_Bits_Cores : Struct
            No_end_in_WP_core01 : Bool := FALSE;
            No_end_in_BP_core01 : Bool := FALSE;
            Always_ON_in_WP_core01 : Bool := TRUE;
            Always_ON_in_BP_core01 : Bool := TRUE;
            Inverted_end_in_WP_core01 : Bool := FALSE;
            Inverted_end_in_BP_core01 : Bool := FALSE;
            No_hydraulic_core01 : Bool := FALSE;
            Upper_tool_core01 : Bool := FALSE;
            No_end_in_WP_core02 : Bool := FALSE;
            No_end_in_BP_core02 : Bool := FALSE;
            Always_ON_in_WP_core02 : Bool := TRUE;
            Always_ON_in_BP_core02 : Bool := TRUE;
            Inverted_end_in_WP_core02 : Bool := FALSE;
            Inverted_end_in_BP_core02 : Bool := FALSE;
            No_hydraulic_core02 : Bool := FALSE;
            Upper_tool_core02 : Bool := FALSE;
            No_end_in_WP_core03 : Bool := FALSE;
            No_end_in_BP_core03 : Bool := FALSE;
            Always_ON_in_WP_core03 : Bool := TRUE;
            Always_ON_in_BP_core03 : Bool := TRUE;
            Inverted_end_in_WP_core03 : Bool := FALSE;
            Inverted_end_in_BP_core03 : Bool := FALSE;
            No_hydraulic_core03 : Bool := FALSE;
            Upper_tool_core03 : Bool := FALSE;
            No_end_in_WP_core04 : Bool := FALSE;
            No_end_in_BP_core04 : Bool := FALSE;
            Always_ON_in_WP_core04 : Bool := TRUE;
            Always_ON_in_BP_core04 : Bool := TRUE;
            Inverted_end_in_WP_core04 : Bool := FALSE;
            Inverted_end_in_BP_core04 : Bool := FALSE;
            No_hydraulic_core04 : Bool := FALSE;
            Upper_tool_core04 : Bool := FALSE;
            No_end_in_WP_core05 : Bool := FALSE;
            No_end_in_BP_core05 : Bool := FALSE;
            Always_ON_in_WP_core05 : Bool := TRUE;
            Always_ON_in_BP_core05 : Bool := TRUE;
            Inverted_end_in_WP_core05 : Bool := FALSE;
            Inverted_end_in_BP_core05 : Bool := TRUE;
            No_hydraulic_core05 : Bool := FALSE;
            Upper_tool_core05 : Bool := FALSE;
            No_end_in_WP_core06 : Bool := FALSE;
            No_end_in_BP_core06 : Bool := FALSE;
            Always_ON_in_WP_core06 : Bool := TRUE;
            Always_ON_in_BP_core06 : Bool := TRUE;
            Inverted_end_in_WP_core06 : Bool := FALSE;
            Inverted_end_in_BP_core06 : Bool := TRUE;
            No_hydraulic_core06 : Bool := FALSE;
            Upper_tool_core06 : Bool := FALSE;
            No_end_in_WP_core07 : Bool := TRUE;
            No_end_in_BP_core07 : Bool := TRUE;
            Always_ON_in_WP_core07 : Bool := TRUE;
            Always_ON_in_BP_core07 : Bool := TRUE;
            Inverted_end_in_WP_core07 : Bool := FALSE;
            Inverted_end_in_BP_core07 : Bool := FALSE;
            No_hydraulic_core07 : Bool := FALSE;
            Upper_tool_core07 : Bool := FALSE;
            No_end_in_WP_core08 : Bool := FALSE;
            No_end_in_BP_core08 : Bool := FALSE;
            Always_ON_in_WP_core08 : Bool := TRUE;
            Always_ON_in_BP_core08 : Bool := TRUE;
            Inverted_end_in_WP_core08 : Bool := FALSE;
            Inverted_end_in_BP_core08 : Bool := TRUE;
            No_hydraulic_core08 : Bool := FALSE;
            Upper_tool_core08 : Bool := FALSE;
            No_end_in_WP_core09 : Bool := FALSE;
            No_end_in_BP_core09 : Bool := FALSE;
            Always_ON_in_WP_core09 : Bool := TRUE;
            Always_ON_in_BP_core09 : Bool := TRUE;
            Inverted_end_in_WP_core09 : Bool := FALSE;
            Inverted_end_in_BP_core09 : Bool := TRUE;
            No_hydraulic_core09 : Bool := FALSE;
            Upper_tool_core09 : Bool := FALSE;
            No_end_in_WP_core10 : Bool := FALSE;
            No_end_in_BP_core10 : Bool := FALSE;
            Always_ON_in_WP_core10 : Bool := TRUE;
            Always_ON_in_BP_core10 : Bool := TRUE;
            Inverted_end_in_WP_core10 : Bool := FALSE;
            Inverted_end_in_BP_core10 : Bool := FALSE;
            No_hydraulic_core10 : Bool := FALSE;
            Upper_tool_core10 : Bool := FALSE;
            No_end_in_WP_core11 : Bool := FALSE;
            No_end_in_BP_core11 : Bool := FALSE;
            Always_ON_in_WP_core11 : Bool := TRUE;
            Always_ON_in_BP_core11 : Bool := TRUE;
            Inverted_end_in_WP_core11 : Bool := FALSE;
            Inverted_end_in_BP_core11 : Bool := FALSE;
            No_hydraulic_core11 : Bool := FALSE;
            Upper_tool_core11 : Bool := FALSE;
            No_end_in_WP_core12 : Bool := FALSE;
            No_end_in_BP_core12 : Bool := FALSE;
            Always_ON_in_WP_core12 : Bool := TRUE;
            Always_ON_in_BP_core12 : Bool := TRUE;
            Inverted_end_in_WP_core12 : Bool := FALSE;
            Inverted_end_in_BP_core12 : Bool := FALSE;
            No_hydraulic_core12 : Bool := FALSE;
            Upper_tool_core12 : Bool := FALSE;
            No_end_in_WP_core13 : Bool := FALSE;
            No_end_in_BP_core13 : Bool := FALSE;
            Always_ON_in_WP_core13 : Bool := TRUE;
            Always_ON_in_BP_core13 : Bool := TRUE;
            Inverted_end_in_WP_core13 : Bool := FALSE;
            Inverted_end_in_BP_core13 : Bool := FALSE;
            No_hydraulic_core13 : Bool := FALSE;
            Upper_tool_core13 : Bool := FALSE;
            No_end_in_WP_core14 : Bool := FALSE;
            No_end_in_BP_core14 : Bool := FALSE;
            Always_ON_in_WP_core14 : Bool := TRUE;
            Always_ON_in_BP_core14 : Bool := TRUE;
            Inverted_end_in_WP_core14 : Bool := FALSE;
            Inverted_end_in_BP_core14 : Bool := FALSE;
            No_hydraulic_core14 : Bool := FALSE;
            Upper_tool_core14 : Bool := FALSE;
            No_end_in_WP_core15 : Bool := FALSE;
            No_end_in_BP_core15 : Bool := FALSE;
            Always_ON_in_WP_core15 : Bool := TRUE;
            Always_ON_in_BP_core15 : Bool := TRUE;
            Inverted_end_in_WP_core15 : Bool := FALSE;
            Inverted_end_in_BP_core15 : Bool := FALSE;
            No_hydraulic_core15 : Bool := FALSE;
            Upper_tool_core15 : Bool := FALSE;
            No_end_in_WP_core16 : Bool := FALSE;
            No_end_in_BP_core16 : Bool := FALSE;
            Always_ON_in_WP_core16 : Bool := TRUE;
            Always_ON_in_BP_core16 : Bool := TRUE;
            Inverted_end_in_WP_core16 : Bool := FALSE;
            Inverted_end_in_BP_core16 : Bool := FALSE;
            No_hydraulic_core16 : Bool := FALSE;
            Upper_tool_core16 : Bool := FALSE;
            No_end_in_WP_core17 : Bool := FALSE;
            No_end_in_BP_core17 : Bool := FALSE;
            Always_ON_in_WP_core17 : Bool := TRUE;
            Always_ON_in_BP_core17 : Bool := TRUE;
            Inverted_end_in_WP_core17 : Bool := FALSE;
            Inverted_end_in_BP_core17 : Bool := FALSE;
            No_hydraulic_core17 : Bool := FALSE;
            Upper_tool_core17 : Bool := FALSE;
            No_end_in_WP_core18 : Bool := FALSE;
            No_end_in_BP_core18 : Bool := FALSE;
            Always_ON_in_WP_core18 : Bool := TRUE;
            Always_ON_in_BP_core18 : Bool := TRUE;
            Inverted_end_in_WP_core18 : Bool := FALSE;
            Inverted_end_in_BP_core18 : Bool := FALSE;
            No_hydraulic_core18 : Bool := FALSE;
            Upper_tool_core18 : Bool := FALSE;
            No_end_in_WP_core19 : Bool := FALSE;
            No_end_in_BP_core19 : Bool := FALSE;
            Always_ON_in_WP_core19 : Bool := TRUE;
            Always_ON_in_BP_core19 : Bool := TRUE;
            Inverted_end_in_WP_core19 : Bool := FALSE;
            Inverted_end_in_BP_core19 : Bool := FALSE;
            No_hydraulic_core19 : Bool := FALSE;
            Upper_tool_core19 : Bool := FALSE;
            No_end_in_WP_core20 : Bool := FALSE;
            No_end_in_BP_core20 : Bool := FALSE;
            Always_ON_in_WP_core20 : Bool := TRUE;
            Always_ON_in_BP_core20 : Bool := TRUE;
            Inverted_end_in_WP_core20 : Bool := FALSE;
            Inverted_end_in_BP_core20 : Bool := FALSE;
            No_hydraulic_core20 : Bool := FALSE;
            Upper_tool_core20 : Bool := FALSE;
            No_end_in_WP_core21 : Bool := FALSE;
            No_end_in_BP_core21 : Bool := FALSE;
            Always_ON_in_WP_core21 : Bool := TRUE;
            Always_ON_in_BP_core21 : Bool := TRUE;
            Inverted_end_in_WP_core21 : Bool := FALSE;
            Inverted_end_in_BP_core21 : Bool := FALSE;
            No_hydraulic_core21 : Bool := FALSE;
            Upper_tool_core21 : Bool := FALSE;
            No_end_in_WP_core22 : Bool := FALSE;
            No_end_in_BP_core22 : Bool := FALSE;
            Always_ON_in_WP_core22 : Bool := TRUE;
            Always_ON_in_BP_core22 : Bool := TRUE;
            Inverted_end_in_WP_core22 : Bool := FALSE;
            Inverted_end_in_BP_core22 : Bool := FALSE;
            No_hydraulic_core22 : Bool := FALSE;
            Upper_tool_core22 : Bool := FALSE;
            No_end_in_WP_core23 : Bool := FALSE;
            No_end_in_BP_core23 : Bool := FALSE;
            Always_ON_in_WP_core23 : Bool := TRUE;
            Always_ON_in_BP_core23 : Bool := TRUE;
            Inverted_end_in_WP_core23 : Bool := FALSE;
            Inverted_end_in_BP_core23 : Bool := FALSE;
            No_hydraulic_core23 : Bool := FALSE;
            Upper_tool_core23 : Bool := FALSE;
            No_end_in_WP_core24 : Bool := FALSE;
            No_end_in_BP_core24 : Bool := FALSE;
            Always_ON_in_WP_core24 : Bool := TRUE;
            Always_ON_in_BP_core24 : Bool := TRUE;
            Inverted_end_in_WP_core24 : Bool := FALSE;
            Inverted_end_in_BP_core24 : Bool := FALSE;
            No_hydraulic_core24 : Bool := FALSE;
            Upper_tool_core24 : Bool := FALSE;
            No_end_in_WP_core25 : Bool := FALSE;
            No_end_in_BP_core25 : Bool := FALSE;
            Always_ON_in_WP_core25 : Bool := TRUE;
            Always_ON_in_BP_core25 : Bool := TRUE;
            Inverted_end_in_WP_core25 : Bool := FALSE;
            Inverted_end_in_BP_core25 : Bool := FALSE;
            No_hydraulic_core25 : Bool := FALSE;
            Upper_tool_core25 : Bool := FALSE;
            No_end_in_WP_core26 : Bool := FALSE;
            No_end_in_BP_core26 : Bool := FALSE;
            Always_ON_in_WP_core26 : Bool := TRUE;
            Always_ON_in_BP_core26 : Bool := TRUE;
            Inverted_end_in_WP_core26 : Bool := FALSE;
            Inverted_end_in_BP_core26 : Bool := FALSE;
            No_hydraulic_core26 : Bool := FALSE;
            Upper_tool_core26 : Bool := FALSE;
            No_end_in_WP_core27 : Bool := FALSE;
            No_end_in_BP_core27 : Bool := FALSE;
            Always_ON_in_WP_core27 : Bool := TRUE;
            Always_ON_in_BP_core27 : Bool := TRUE;
            Inverted_end_in_WP_core27 : Bool := FALSE;
            Inverted_end_in_BP_core27 : Bool := FALSE;
            No_hydraulic_core27 : Bool := FALSE;
            Upper_tool_core27 : Bool := FALSE;
            No_end_in_WP_core28 : Bool := FALSE;
            No_end_in_BP_core28 : Bool := FALSE;
            Always_ON_in_WP_core28 : Bool := TRUE;
            Always_ON_in_BP_core28 : Bool := TRUE;
            Inverted_end_in_WP_core28 : Bool := FALSE;
            Inverted_end_in_BP_core28 : Bool := FALSE;
            No_hydraulic_core28 : Bool := FALSE;
            Upper_tool_core28 : Bool := FALSE;
            No_end_in_WP_core29 : Bool := FALSE;
            No_end_in_BP_core29 : Bool := FALSE;
            Always_ON_in_WP_core29 : Bool := TRUE;
            Always_ON_in_BP_core29 : Bool := TRUE;
            Inverted_end_in_WP_core29 : Bool := FALSE;
            Inverted_end_in_BP_core29 : Bool := FALSE;
            No_hydraulic_core29 : Bool := FALSE;
            Upper_tool_core29 : Bool := FALSE;
            No_end_in_WP_core30 : Bool := FALSE;
            No_end_in_BP_core30 : Bool := FALSE;
            Always_ON_in_WP_core30 : Bool := TRUE;
            Always_ON_in_BP_core30 : Bool := TRUE;
            Inverted_end_in_WP_core30 : Bool := FALSE;
            Inverted_end_in_BP_core30 : Bool := FALSE;
            No_hydraulic_core30 : Bool := FALSE;
            Upper_tool_core30 : Bool := FALSE;
            No_end_in_WP_core31 : Bool := FALSE;
            No_end_in_BP_core31 : Bool := FALSE;
            Always_ON_in_WP_core31 : Bool := TRUE;
            Always_ON_in_BP_core31 : Bool := TRUE;
            Inverted_end_in_WP_core31 : Bool := FALSE;
            Inverted_end_in_BP_core31 : Bool := FALSE;
            No_hydraulic_core31 : Bool := FALSE;
            Upper_tool_core31 : Bool := FALSE;
            No_end_in_WP_core32 : Bool := FALSE;
            No_end_in_BP_core32 : Bool := FALSE;
            Always_ON_in_WP_core32 : Bool := TRUE;
            Always_ON_in_BP_core32 : Bool := TRUE;
            Inverted_end_in_WP_core32 : Bool := FALSE;
            Inverted_end_in_BP_core32 : Bool := FALSE;
            No_hydraulic_core32 : Bool := FALSE;
            Upper_tool_core32 : Bool := FALSE;
         END_STRUCT;
         Special_Bits : Struct
            Spare_0_0 : Bool := FALSE;